SwitchIO70313.xExitEnable:=(ConveyorIO70199.xEmpty AND (ConveyorIO70152.diDesConveyor=70199 OR ConveyorIO70152.diDesConveyor=70154))
													OR (ConveyorIO701100.xEmpty AND (ConveyorIO70152.diDesConveyor=701100 OR ConveyorIO70152.diDesConveyor=70155));
ConveyorIO70192.xUnloadCCW:=ConveyorIO70192.diDesConveyor=701100 OR ConveyorIO70192.diDesConveyor=70155;
ConveyorIO70199.xLoad:=ConveyorIO70192.xNextRun AND (ConveyorIO70152.diDesConveyor=70199 OR ConveyorIO70152.diDesConveyor=70154);
ConveyorIO70199.xUnload:=ConveyorIO70154.xEmpty AND ConveyorIO70199.diDesConveyor=70154;
ConveyorIO70154.xLoad:=ConveyorIO70199.xNextRun;
m_xtonConveyor70199Reset(IN:=NOT ConveyorIO70199.xCWPresent,PT:=T#10s ,Q:= ConveyorIO70199.xPutInto,ET:= m_xtonConveyor70199CurTime );
m_xtonConveyor70154Reset(IN:=NOT ConveyorIO70154.xCWPresent,PT:=T#10s ,Q:= ConveyorIO70154.xPutInto,ET:= m_xtonConveyor70154CurTime );
ConveyorIO701100.xLoad:=ConveyorIO70192.xNextRun AND (ConveyorIO70152.diDesConveyor=701100 OR ConveyorIO70152.diDesConveyor=70155);
ConveyorIO701100.xUnload:=ConveyorIO70155.xEmpty AND ConveyorIO701100.diDesConveyor=70155;
ConveyorIO70155.xLoad:=ConveyorIO701100.xNextRun;
m_xtonConveyor701100Reset(IN:=NOT ConveyorIO701100.xCWPresent,PT:=T#10s ,Q:= ConveyorIO701100.xPutInto,ET:=m_xtonConveyor701100CurTime );
m_xtonConveyor70155Reset(IN:=NOT ConveyorIO70155.xCWPresent,PT:=T#10s ,Q:= ConveyorIO70155.xPutInto,ET:= m_xtonConveyor70155CurTime);



(*3#下层入库*)
(*
IF  ConveyorIO70160.xLoad
	THEN Y2C6:=1;
END_IF;
IF NOT  ConveyorIO70160.xEmpty
	THEN  Y2C6:=0;
END_IF;*)
switch70315(ConveyorEntryIO:= ConveyorIO70160 ,ConveyorExitIO:= ConveyorIO70194 ,SwitchIO:= SwitchIO70315);
SwitchIO70315.xLiftCylinderExtendInit:=1;
SwitchIO70315.xSwithEnable:=1;
Y2C6:=SwitchIO70315.xLiftCylinderExtend;
SwitchIO70315.xLiftCylinderExtendDetect:=XDA;
SwitchIO70315.xLiftCylinderRetractDetect:=XDB;

SwitchIO70315.xExitEnable:=(ConveyorIO701103.xEmpty AND (ConveyorIO70160.diDesConveyor=701103 OR ConveyorIO70160.diDesConveyor=70162))
													OR (ConveyorIO701104.xEmpty AND (ConveyorIO70160.diDesConveyor=701104 OR ConveyorIO70160.diDesConveyor=70163));
ConveyorIO70194.xUnloadCCW:=ConveyorIO70194.diDesConveyor=701103 OR ConveyorIO70194.diDesConveyor=70162;
ConveyorIO701103.xLoad:=ConveyorIO70194.xNextRun AND (ConveyorIO70160.diDesConveyor=701103 OR ConveyorIO70160.diDesConveyor=70162);
ConveyorIO701103.xUnload:=ConveyorIO70162.xEmpty AND ConveyorIO701103.diDesConveyor=70162;
ConveyorIO70162.xLoad:=ConveyorIO701103.xNextRun;
m_xtonConveyor701103Reset(IN:=NOT ConveyorIO701103.xCWPresent,PT:=T#10s ,Q:= ConveyorIO701103.xPutInto,ET:= m_xtonConveyor701103CurTime );
m_xtonConveyor70162Reset(IN:=NOT ConveyorIO70162.xCWPresent,PT:=T#10s ,Q:= ConveyorIO70162.xPutInto,ET:= m_xtonConveyor70162CurTime );
ConveyorIO701104.xLoad:=ConveyorIO70194.xNextRun AND (ConveyorIO70160.diDesConveyor=701104 OR ConveyorIO70160.diDesConveyor=70163);
ConveyorIO701104.xUnload:=ConveyorIO70163.xEmpty AND ConveyorIO701104.diDesConveyor=70163;
ConveyorIO70163.xLoad:=ConveyorIO701104.xNextRun;
m_xtonConveyor701104Reset(IN:=NOT ConveyorIO701104.xCWPresent,PT:=T#10s ,Q:= ConveyorIO701104.xPutInto,ET:=m_xtonConveyor701104CurTime );
m_xtonConveyor70163Reset(IN:=NOT ConveyorIO70163.xCWPresent,PT:=T#10s ,Q:= ConveyorIO70163.xPutInto,ET:= m_xtonConveyor70163CurTime);


(*2，3#下层出库,只写了3#的*)
(*23出库任务抢占*)
	m_Task70314(xCondition:= m_Task70314Condition ,
							xTaskComplete:=LDP(TRUE,ConveyorIO70193.xEmpty) ,
							xReset:= g_xResetSingle AND g_diDeviceIDSelect=70193 ,
							iPriority:= m_iTask70314  );
		m_Task70314Condition[1]:=NOT ConveyorIO701101.xEmpty;
		m_Task70314Condition[2]:=NOT ConveyorIO701102.xEmpty;
		
m_xtonConveyor70159Reset(IN:= ConveyorIO70159.xCWPresent,PT:=T#10s ,Q:= ConveyorIO70159.xPutInto,ET:= m_xtonConveyor70159CurTime );
m_xtonConveyor701102Reset(IN:= ConveyorIO701102.xCWPresent,PT:=T#10s ,Q:= ConveyorIO701102.xPutInto,ET:= m_xtonConveyor701102CurTime );
ConveyorIO70159.xUnload:=ConveyorIO701102.xEmpty;
ConveyorIO701102.xLoad:=ConveyorIO70159.xNextRun;
ConveyorIO701102.xUnload:=ConveyorIO70193.xEmpty AND m_iTask70314=2;

m_xtonConveyor70158Reset(IN:= ConveyorIO70158.xCWPresent,PT:=T#10s ,Q:= ConveyorIO70158.xPutInto,ET:= m_xtonConveyor70158CurTime );
m_xtonConveyor701101Reset(IN:= ConveyorIO701101.xCWPresent,PT:=T#10s ,Q:= ConveyorIO701101.xPutInto,ET:= m_xtonConveyor701101CurTime );
ConveyorIO70158.xUnload:=ConveyorIO701101.xEmpty;
ConveyorIO701101.xLoad:=ConveyorIO70158.xNextRun;
ConveyorIO701101.xUnload:=ConveyorIO70193.xEmpty AND m_iTask70314=1;

ConveyorIO70193.xLoad:=ConveyorIO701102.xNextRun OR ConveyorIO701101.xNextRun;
ConveyorIO70193.xloadCCW:=ConveyorIO701102.xNextRun;
IF  NOT ConveyorIO70193.xEmpty
	THEN Y2C4:=1;(*193转去156顶升*)
END_IF;
ConveyorIO70156.xLoad:= NOT ConveyorIO70193.xEmpty ;
IF NOT  ConveyorIO70156.xEmpty
	THEN 
	Y2C4:=0;
END_IF;
m_xtonConveyor70156Reset(IN:=NOT ConveyorIO70156.xCWPresent,PT:=T#10s ,Q:= ConveyorIO70156.xPutInto,ET:= m_xtonConveyor70156CurTime );
Y33B:=ConveyorIO701102.xNextRun;(*3#出库阻挡*)
Y33A:=ConveyorIO701101.xNextRun;(*2#出库阻挡*)
ConveyorIO70193.xPutInto:=NOT  ConveyorIO70156.xEmpty;
(*最靠近电柜那个出库线体*)
switch70327(ConveyorEntryIO:=ConveyorIO701118,ConveyorExitIO:= ConveyorIO701116_1 ,SwitchIO:= SwitchIO70327);
Y2DE:=SwitchIO70327.xLiftCylinderExtend;
SwitchIO70327.xLiftCylinderExtendDetect:=X155;
SwitchIO70327.xLiftCylinderRetractDetect:=X156;

Conveyor701116_1(ConveyorMotor:= ConveyorIO701116_1 );
ConveyorIO701116_1.xCWPresent:=ConveyorIO701118.xCWPresent;

m_xtonConveyor701120Reset(IN:=ConveyorIO701120.xCWPresent,PT:=T#10s ,Q:= ConveyorIO701120.xPutInto,ET:= m_xtonConveyor701120CurTime );
m_xtonConveyor701119Reset(IN:=ConveyorIO701119.xCWPresent,PT:=T#10s ,Q:= ConveyorIO701119.xPutInto,ET:= m_xtonConveyor701119CurTime );
ConveyorIO701119.tLoadDelay:=t#3s;
ConveyorIO701120.xUnload:=ConveyorIO701119.xEmpty;
ConveyorIO701119.xLoad:=ConveyorIO701120.xNextRun;
ConveyorIO701119.xUnload:=ConveyorIO701118.xEmpty;
SwitchIO70327.xEntryEnable:=ConveyorIO701119.xNextRun;
SwitchIO70327.xSwithEnable:=1;
SwitchIO70327.xExitEnable:=ConveyorIO701116.xEmpty;
ConveyorIO701116.xLoad:=ConveyorIO701116_1.xNextRun;

(*回流部分去分容线体*)
ConveyorIO70141.xLoad:=X3D;
Y2BA:=ConveyorIO70141.xEmpty;
m_xtonConveyor70141Reset(IN:=NOT ConveyorIO70141.xCWPresent,PT:=T#8s ,Q:= ConveyorIO70141.xPutInto,ET:= m_xtonConveyor70141CurTime );

(*————————上层空框回流————————————*)
ConveyorIO70134.xUnload:=ConveyorIO70133.xEmpty;
ConveyorIO70133.xLoad:=ConveyorIO70134.xNextRun;
ConveyorIO70133.xUnload:=ConveyorIO70132.xEmpty;
ConveyorIO70132.xLoad:=ConveyorIO70133.xNextRun;
ConveyorIO70132.xUnload:=ConveyorIO70131.xEmpty;
ConveyorIO70131.xLoad:=ConveyorIO70132.xNextRun;
ConveyorIO70131.xUnload:=ConveyorIO70130.xEmpty;
ConveyorIO70130.xLoad:=ConveyorIO70131.xNextRun;
ConveyorIO70130.xUnload:=ConveyorIO70124.xEmpty;
ConveyorIO70124.xLoad:=ConveyorIO70130.xNextRun;
ConveyorIO70124.xUnload:=ConveyorIO70123.xEmpty;
ConveyorIO70123.xLoad:=ConveyorIO70124.xNextRun;
ConveyorIO70123.xUnload:=ConveyorIO70122.xEmpty;
ConveyorIO70122.xLoad:=ConveyorIO70123.xNextRun;
ConveyorIO70122.xUnload:=ConveyorIO70116.xEmpty;
ConveyorIO70116.xLoad:=ConveyorIO70122.xNextRun;
ConveyorIO70116.xUnload:=ConveyorIO70115.xEmpty;
ConveyorIO70115.xLoad:=ConveyorIO70116.xNextRun;
ConveyorIO70115.xUnload:=ConveyorIO70114.xEmpty;
ConveyorIO70114.xLoad:=ConveyorIO70115.xNextRun;
ConveyorIO70114.xUnload:=ConveyorIO70108.xEmpty;
ConveyorIO70108.xLoad:=ConveyorIO70114.xNextRun;
ConveyorIO70108.xUnload:=ConveyorIO70107.xEmpty AND LifterIO70208.iCurrentPos=2; 
(*提升机2*)
LifterIO70208.xMDIExe:=NOT (ConveyorIO70108.xError OR ConveyorIO70142.xError OR ConveyorIO70107.xError);
IF ConveyorIO70107.xEmpty THEN
	LifterIO70208.iDestinationPos:=2;
ELSE
	LifterIO70208.iDestinationPos:=1;
END_IF;
ConveyorIO70107.xLoad:=ConveyorIO70108.xNextRun AND LifterIO70208.iCurrentPos=2;
ConveyorIO70107.xUnload:=ConveyorIO70142.xEmpty AND  LifterIO70208.iCurrentPos=1;
ConveyorIO70142.xLoad:=ConveyorIO70107.xNextRun AND   LifterIO70208.iCurrentPos=1;







(*临时程序,输送出去,不进2号OCV2，不分拣*) 
(*ConveyorIO70166.xUnload:=ConveyorIO70167.xEmpty;*)
(*临时程序,分拣前顶升移载前*)
(*SwitchIO70319.xEntryEnable:=ConveyorIO70166.xNextRun;*)
(*SwitchIO70319.xSwithEnable:=0;*)(*临时程序不分拣*)
(*SwitchIO70319.xExitEnable:=ConveyorIO70169.xEmpty;
SwitchIO70320.xEntryEnable:=ConveyorIO70167.xNextRun;
SwitchIO70320.xSwithEnable:=1;
SwitchIO70320.xExitEnable:=0;*)(*RGV接料处*)


IF g_xAuto AND NOT g_xRGVTcpFailed THEN
	D201:=m_iRGVDestinationPos;
	D202.0:=g_xRGVRemoteAuto;
	D202.1:=(*ConveyorIO70140.xEmpty*)NOT FolderIO70201.o_xExitPremit;(*更换成叠盘机允许下料信号，RGV生成任务*)
	D202.2:=ConveyorIO701111.xEmpty;
	D202.3:=ConveyorIO70144.xEmpty;
	D202.4:=ConveyorIO70148.xEmpty;
	D202.5:=ConveyorIO70152.xEmpty;
	D202.6:=ConveyorIO70156.xEmpty;
	D202.7:=ConveyorIO70160.xEmpty;
	D202.8:=ConveyorIO70164.xEmpty;
	D202.9:=ConveyorIO70170.xEmpty;
	D202.A:=ConveyorIO70174.xEmpty;
	D202.B:=ConveyorIO701116.xEmpty;
	D203.0:=m_xRGVReset;
	D203.1:=ConveyorIO70140.xNextRun;
	D203.2:=ConveyorIO701111.xNextRun;
	D203.3:=ConveyorIO70148.xNextRun;
	D203.4:=ConveyorIO70156.xNextRun;
	D203.5:=ConveyorIO70170.xNextRun;
	D203.6:=ConveyorIO701116.xNextRun;
	D203.A:=g_SemiStart;
	m_iRGVCurrentPos:=D401;
	m_xRGVPositionArrive:=D401.0;
	m_xRGVConveyorEmpty:=D401.1;
	m_xRGVConveyorNextRun:=D402.2;
	ConveyorIO70140.xUnload:=D402.3;
	ConveyorIO701111.xUnload:=D402.4;
	ConveyorIO70144.xLoad:=D402.5;
	ConveyorIO70148.xUnload:=D402.6;
	ConveyorIO70152.xLoad:=D402.7;
	ConveyorIO70156.xUnload:=D402.8;
	ConveyorIO70160.xLoad:=D402.9;
	ConveyorIO70164.xLoad:=D402.A;
	ConveyorIO70170.xUnload:=D402.B;
	ConveyorIO70174.xLoad:=D402.C;
	ConveyorIO701116.xUnload:=D402.D;
	m_xRGVAlarm:=D403.0;
ELSE
	D201:=0;
	D202:=0;
	D203.0:=0;
	D203.1:=0;
	D203.2:=0;
	D203.3:=0;
	D203.4:=0;
	D203.5:=0;
	ConveyorIO70140.xUnload:=0;
	ConveyorIO701111.xUnload:=0;
	ConveyorIO70144.xLoad:=0;
	ConveyorIO70148.xUnload:=0;
	ConveyorIO70152.xLoad:=0;
	ConveyorIO70156.xUnload:=0;
	ConveyorIO70160.xLoad:=0;
	ConveyorIO70164.xLoad:=0;
	ConveyorIO70170.xUnload:=0;
	ConveyorIO70174.xLoad:=0;
END_IF;
g_xAlarm:=ComConveyorIO70104.i_iResponsPCPLC=101;
END_PROGRAM

FUNCTION_BLOCK PreemptivePriority
VAR_INPUT
  xCondition : ARRAY [1..13] OF BOOL;  (* 条件1 *)
  xTaskComplete : BOOL;  (* 任务完成 *)
  xReset : BOOL;  (* 复位 *)
END_VAR
VAR
  xOccupy : BOOL;  (* 占用 *)
END_VAR
VAR_OUTPUT
  iPriority : INT;  (* 输出任务号 *)
END_VAR
VAR
  m_tonConditionDelay : TON;
  m_xConditionDelay : BOOL;
  m_tConditionCurrentTime : TIME;
  m_iLastTask : INT;  (* 上次执行的任务 *)
  m_tpLastTaskPulse1 : TP;
  m_tpLastTaskPulse2 : TP;
  m_tpLastTaskPulse3 : TP;
  m_tpLastTaskPulse4 : TP;
  m_tpLastTaskPulse5 : TP;
  m_xLastTaskPulse : ARRAY [1..13] OF BOOL;
  m_tLastTaskPulse : ARRAY [1..13] OF TIME := [13(T#0s)];
  m_tpLastTaskPulse6 : TON;
  ii : INT;
END_VAR
VAR CONSTANT
  CONDITION_QUANTITY : INT := 9;
END_VAR
VAR
  m_tpLastTaskPulse7 : TON;
  m_tpLastTaskPulse8 : TON;
  m_tpLastTaskPulse9 : TON;
  m_tpLastTaskPulse10 : TON;
  m_tpLastTaskPulse11 : TON;
  m_tpLastTaskPulse12 : TON;
  m_tpLastTaskPulse13 : TON;
END_VAR
(*抢占式优先级块
现在满足13个条件的任务进行抢占式优先级排列
条件满足后延时两秒，开始执行任务，
同一任务连续执行优先级下降
需要改造成任意多个
使用于一个入口多个出口的程序，使用抢占式优先级块
*)
IF LDP(TRUE, xTaskComplete) THEN
	xOccupy:=0;
	iPriority:=0;
END_IF;
(*//任务滤波，延时两秒*)
m_tonConditionDelay(IN:=( xCondition[1]
 	OR xCondition[2]
 	OR xCondition[3]
 	OR xCondition[4]
 	OR xCondition[5]
 	OR xCondition[6]
 	OR xCondition[7]
 	OR xCondition[8]
 	OR xCondition[9]
 	OR xCondition[10]
 	OR xCondition[11]
 	OR xCondition[12]
 	OR xCondition[13]
 	)
 	AND iPriority=0,
 PT:= T#1s,
 Q:= m_xConditionDelay ,
 ET:= m_tConditionCurrentTime );		
(*//判断优先级，上个任务与本次任务相同，延时一秒执行*)
m_tpLastTaskPulse1(IN:= xCondition[1]  AND m_iLastTask=1 AND m_xConditionDelay  ,PT:= T#1s,Q:= m_xLastTaskPulse[1],ET:= m_tLastTaskPulse[1] );
m_tpLastTaskPulse2(IN:= xCondition[2]  AND m_iLastTask=2 AND m_xConditionDelay  ,PT:= T#1s,Q:= m_xLastTaskPulse[2],ET:= m_tLastTaskPulse[2] );
m_tpLastTaskPulse3(IN:= xCondition[3]  AND m_iLastTask=3 AND m_xConditionDelay  ,PT:= T#1s,Q:= m_xLastTaskPulse[3],ET:= m_tLastTaskPulse[3] );
m_tpLastTaskPulse4(IN:= xCondition[4]  AND m_iLastTask=4 AND m_xConditionDelay  ,PT:= T#1s,Q:= m_xLastTaskPulse[4],ET:= m_tLastTaskPulse[4] );
m_tpLastTaskPulse5(IN:= xCondition[5]  AND m_iLastTask=5 AND m_xConditionDelay  ,PT:= T#1s,Q:= m_xLastTaskPulse[5],ET:= m_tLastTaskPulse[5] );
m_tpLastTaskPulse6(IN:= xCondition[6]  AND m_iLastTask=6 AND m_xConditionDelay  ,PT:= T#1s,Q:= m_xLastTaskPulse[6],ET:= m_tLastTaskPulse[6] );
m_tpLastTaskPulse7(IN:= xCondition[7]  AND m_iLastTask=7 AND m_xConditionDelay  ,PT:= T#1s,Q:= m_xLastTaskPulse[7],ET:= m_tLastTaskPulse[7] );
m_tpLastTaskPulse8(IN:= xCondition[8]  AND m_iLastTask=8 AND m_xConditionDelay  ,PT:= T#1s,Q:= m_xLastTaskPulse[8],ET:= m_tLastTaskPulse[8] );
m_tpLastTaskPulse9(IN:= xCondition[9]  AND m_iLastTask=9 AND m_xConditionDelay  ,PT:= T#1s,Q:= m_xLastTaskPulse[9],ET:= m_tLastTaskPulse[9] );
m_tpLastTaskPulse10(IN:= xCondition[10]  AND m_iLastTask=10 AND m_xConditionDelay  ,PT:= T#1s,Q:= m_xLastTaskPulse[10],ET:= m_tLastTaskPulse[10] );
m_tpLastTaskPulse11(IN:= xCondition[11]  AND m_iLastTask=11 AND m_xConditionDelay  ,PT:= T#1s,Q:= m_xLastTaskPulse[11],ET:= m_tLastTaskPulse[11] );
m_tpLastTaskPulse12(IN:= xCondition[12]  AND m_iLastTask=12 AND m_xConditionDelay  ,PT:= T#1s,Q:= m_xLastTaskPulse[12],ET:= m_tLastTaskPulse[12] );
m_tpLastTaskPulse13(IN:= xCondition[13]  AND m_iLastTask=13 AND m_xConditionDelay  ,PT:= T#1s,Q:= m_xLastTaskPulse[13],ET:= m_tLastTaskPulse[13] );
(*//执行*)
FOR ii:=1 TO CONDITION_QUANTITY BY 1 DO 
	IF NOT xCondition[ii] AND NOT xOccupy THEN
		iPriority:=0;
	END_IF;
	IF xCondition[ii] AND NOT xOccupy AND m_xConditionDelay AND NOT  m_xLastTaskPulse[ii]  THEN
		iPriority:=ii;
		xOccupy:=1;
		m_iLastTask:=ii;
	END_IF;
END_FOR;        
(*//复位*)
IF xReset THEN
	iPriority:=0;
	xOccupy:=0;
	m_iLastTask:=0;	
END_IF;
(*//清除占用*)
IF iPriority=0 THEN
	xOccupy:=0;
END_IF;
END_FUNCTION_BLOCK

FUNCTION_BLOCK PriorityQueue
VAR_INPUT
  arrxCondition : ARRAY [1..13] OF QueueElement;
  xTaskComplete : BOOL;  (* 任务完成 *)
  xReset : BOOL;  (* 复位 *)
END_VAR
VAR
  xOccupy : BOOL;  (* 占用 *)
END_VAR
VAR_OUTPUT
  iPriority : INT;  (* 输出任务号 *)
END_VAR
VAR
  jj : INT;
END_VAR
VAR CONSTANT
  CONDITION_QUANTITY : INT := 9;
END_VAR
VAR_IN_OUT
  arriTaskStack : ARRAY [0..13] OF INT;
END_VAR
VAR
  ii : INT;
  kk : INT;
  arrxConditionDelay : ARRAY [1..13] OF BOOL;
  arrxConditionEdgeDetect : ARRAY [1..13] OF BOOL;
  arrxDelayEdgeDetect : ARRAY [1..13] OF BOOL;
  arriDelayCounter : ARRAY [1..13] OF INT;
  ll : INT;
  Temp : INT;
  mm : INT;
  nn : INT;
  Temp2 : INT;
  oo : INT;
END_VAR
(****************************************************************************)
(*
一般情况多对一的任务调度采用这个结构，排队通过出口
优先级功能块，存储任意条件的优先级，实现栈功能先入先出，
复位功能还有问题，
出入栈式优先级块，满足条件后入栈，先入先出，在栈尾加载新任务
栈首为当前执行的任务，任务完成使用上升沿触发，触发后栈首元素弹出

复位功能清空堆栈，栈的容量在CONDITION_QUANTITY 设置
增加了结构体，结构体中带有一个条件函数，和一个优先级指示
任务完成后通过凭借优先级来排序，优先级高的条件先执行   优先级排序是从小到大的，数值小的优先级高
防止干扰，增加了任务的1秒的延时
*)

(***************************************************************************)
(*(//入栈*)
FOR ii:=1 TO CONDITION_QUANTITY BY 1 DO
	(*//循环内无法用定时器，改用计数器的形式*)
	IF arrxCondition[ii].xCondition AND SM411 (*//0.2秒的方波信号，如果移植需要修改成两个定时器*)
		AND arriDelayCounter[ii]<6  (* //计数为6，5个0.2秒的方波，所以为1秒*)
		AND NOT arrxDelayEdgeDetect[ii] THEN    (*//循环内无法用沿函数，增加锁定标志位*)
		arriDelayCounter[ii]:=arriDelayCounter[ii]+1;   (*//计数*)
	END_IF;
	IF NOT arrxCondition[ii].xCondition THEN
		arriDelayCounter[ii]:=0;   (*//计数清零*)
	END_IF;
	arrxDelayEdgeDetect[ii]:=arrxCondition[ii].xCondition AND SM411;  (*//沿函数锁*)
	IF arriDelayCounter[ii]=5 AND NOT arrxConditionEdgeDetect[ii] THEN;  (*//条件满足1秒后*)
		FOR kk:=0 TO CONDITION_QUANTITY BY 1 DO    
			IF arriTaskStack[kk]=0 THEN
				arriTaskStack[kk]:=ii;   (*//栈尾添加*)
				EXIT;
			END_IF;		
		END_FOR;
	END_IF;	
	arrxConditionEdgeDetect[ii]:=arriDelayCounter[ii]=5;  (*//边沿*)
END_FOR;
(*//栈顶任务为当前执行的任务**)
iPriority:=arriTaskStack[0]; 
(*//栈顶任务完成，弹出*)
IF 	LDP(TRUE, xTaskComplete) THEN
	FOR jj:=0 TO CONDITION_QUANTITY-1 BY 1 DO
		arriTaskStack[jj]:=arriTaskStack[jj+1];
	END_FOR;
	arriTaskStack[CONDITION_QUANTITY]:=0;(*//栈尾清零*)
	(*//排序，使用插入排序*)
	FOR oo:=0 TO CONDITION_QUANTITY BY 1 DO
		IF arriTaskStack[oo]=0 THEN
			EXIT;  (* //寻找栈中不为零的元素  ，防止0元素进入条件查找的时候报错*)
		END_IF;
	END_FOR;
	(*//插入排序insertionsort*)
	FOR mm:=1 TO oo-1  BY 1 DO   (*//从1开始*)
		Temp:=arriTaskStack[mm];  (*//当前数据记录 *)
		Temp2:=arrxCondition[arriTaskStack[mm]].iPriority;  (*//当前优先级记录 *)
		nn:=mm;  (*//指针赋值*)
		WHILE  (nn>0 AND Temp2< arrxCondition[arriTaskStack[nn-1]].iPriority)  DO  (*//优先级比较，当前优先级小于他前面元素优先级的时候*)
			 arriTaskStack[nn] := arriTaskStack[nn-1] ;  (*//优先级低的向后复制，比TEMP2大的元素都要复制到下一个位置*)
			 nn:=nn-1;
		END_WHILE;
		arriTaskStack[nn]:=Temp; (*//把当前数据放在合适的位置*)
	END_FOR;
END_IF;
(*//复位*)
IF xReset THEN
	FOR jj:=0 TO CONDITION_QUANTITY BY 1 DO
		arriTaskStack[jj]:=0;
	END_FOR;
	FOR ll:=1 TO CONDITION_QUANTITY BY 1 DO
		arrxConditionEdgeDetect[ll]:=0;
		arriDelayCounter[ll]:=0;
	END_FOR;
END_IF;
END_FUNCTION_BLOCK

FUNCTION_BLOCK Servo
Y380:=1;
END_FUNCTION_BLOCK

FUNCTION_BLOCK ShuttleCar
VAR_IN_OUT
  ShuttleCarInOut : ShuttleCarIO;
END_VAR
VAR
  m_tonBrakeDelay : TON;  (* 延时 *)
  m_tBrakeDelayCurrentTime : TIME;
  m_tonArriveDelay : TON;  (* 到达延时计时器 *)
  m_xArriveDelay : BOOL;  (* 到达延时 *)
  m_tArriveDelayCurrentTime : TIME;  (* 到达延时当前时间 *)
  m_xInit : BOOL;  (* 初始化标志位 *)
  m_tonPauseDelay : TON;  (* 暂停减速 *)
  m_tPauseDelayCurrentTime : TIME;  (* 暂停延时当前时间 *)
  m_tonOvertimeAlarm : TON;  (* 超时报警定时器 *)
  m_tOvertimeCurrentTime : TIME;  (* 超时报警当前时间 *)
END_VAR
(*******************************************************************
输送小车程序，可用于使用认址片控制位置的输送车程序，可用于控制提升机，
使用了限位捕捉程序防止小车惯性过大冲过限位后继续行走，捕捉程序采用反
转复位，这样设计有弊端可能反转复位后车的位置并没有回到限位以内,当两个
限位同时碰到的时候，会使运料小车进入死锁状态，通过xPassLimit来解开死锁，
可以在触摸屏中使用一个带权限的按钮来进行控制，配合ShuttleCarCurrentPos
函数来计算位置信息
增加自动开始后将当前位置置为零的信号防止设备停在两个位置开关的中间
修改信息  修改后请增加版本
2018-1-22增加到位延时：到位延时时间可以设置，适应双向到位的位置开关，通过调整延时时间让穿梭车停在到位开关的中间
增加气缸控制信号 ShuttleCarInOut.xCylinder
增加抱闸延时 ShuttleCarInOut.tBrakeDelay
增加超时报警 ShuttleCarInOut.xOvertimeAlarm
YAO      V1.0
2018-1-22 YAO V1.1
2018-6-3：增加点动xMoveStep，单体报警复位
接口说明：
输入：
xReady    准备就绪信号，接变频器的准备就绪，无准备就绪信号的设备常置1
xForward   手动 正转
xBackward 手动 反转
iCurrentPos 当前位置信息，由外部函数给出
iDestinationPos  目标位置，自动情况下判断目标位置和当前位置的差，选择前进或后退
xPosLimit 正方向限位  常闭信号
xNegLimit 反方向限位  常闭信号
xMDIExe   自动行走使能
xPassLimit 限位屏蔽
tArriveDelay 到位延时时间设置，当前位置等于目标位置后延时相应时间后停止，默认为0
xCylinder 如果是气缸的把这个标志位置为1，
tBrakeDelay 打开抱闸延时，默认100ms。行走后会延时相应的时间打开抱闸，防止提升轴的掉落
xLooseDetect 松绳检测开关
输出：
xCW 正转输出
xCCW 反转输出
xBrake 抱闸输出 
xMDIDone 自动行走完成信号
xPosLimitCatch 正限位报警
xNegLimitCatch 负限位报警
xBusy 工作中信号
xLooseAlarm 松绳报警，报警后不可以下降，提升后如果没有松绳检测开关后复位报警信号


********************************************************************)
IF NOT m_xInit THEN
	ShuttleCarInOut.tArriveDelay:=T#0s;   (*到位延时初始化为0*)
	ShuttleCarInOut.tBrakeDelay:=T#100ms;(*抱闸延时初始化为100ms*)
	ShuttleCarInOut.tSetOverTime:=T#60s;(*超时报警初始化为1分钟*)
	m_xInit:=1;
END_IF;
(*如果是气缸的话屏蔽限位和Ready信号*)
IF ShuttleCarInOut.xCylinder THEN
	ShuttleCarInOut.xPosLimit:=1;
	ShuttleCarInOut.xNegLimit:=1;
	ShuttleCarInOut.xReady:=1;
END_IF;
(*限位捕捉，防止冲过限位开关，反转后复位*)
ShuttleCarInOut.xPosLimitCatch:=LDF(TRUE,ShuttleCarInOut.xPosLimit) OR ShuttleCarInOut.xPosLimitCatch;
IF ShuttleCarInOut.xCCW THEN  
	ShuttleCarInOut.xPosLimitCatch:=0;
END_IF;

ShuttleCarInOut.xNegLimitCatch:=LDF(TRUE,ShuttleCarInOut.xNegLimit) OR ShuttleCarInOut.xNegLimitCatch;
(*松绳报警*)
IF LDP(TRUE,ShuttleCarInOut.xLooseDetect) THEN	
	ShuttleCarInOut.xLooseAlarm:=1;
END_IF;
(*提升复位报警*)
IF ShuttleCarInOut.xCW AND NOT  ShuttleCarInOut.xLooseDetect THEN   
	ShuttleCarInOut.xLooseAlarm:=0; 
END_IF;

IF ShuttleCarInOut.xCW THEN   
	ShuttleCarInOut.xNegLimitCatch:=0; 
END_IF;

IF ShuttleCarInOut.xPassLimit OR
	g_xReset OR   (*增加复位按钮*)
	(ShuttleCarInOut.xNegLimitCatch 
	AND ShuttleCarInOut.xPosLimitCatch)  THEN  
	ShuttleCarInOut.xNegLimitCatch:=0; 
	ShuttleCarInOut.xPosLimitCatch:=0;
	ShuttleCarInOut.xLooseAlarm:=0;
END_IF;
IF ShuttleCarInOut.xReady AND g_xEStop THEN
(*手动*)
    IF g_xManual THEN  
	    IF ShuttleCarInOut.xForward 
			AND ShuttleCarInOut.xBackward=0 
			AND ShuttleCarInOut.xCCW=0 
			AND ShuttleCarInOut.xPosLimitCatch=0  THEN
		    ShuttleCarInOut.xCW:=1;
		    ELSE
		    ShuttleCarInOut.xCW:=0;
	    END_IF;
	    IF ShuttleCarInOut.xBackward 
			AND ShuttleCarInOut.xForward=0 
			AND ShuttleCarInOut.xCW=0 
			AND ShuttleCarInOut.xNegLimitCatch=0 
			AND ShuttleCarInOut.xLooseAlarm=0
			AND G_xEStop THEN  
		    ShuttleCarInOut.xCCW:=1;
		    ELSE
		    ShuttleCarInOut.xCCW:=0;
	    END_IF;
    END_IF;
    (**********)
(*自动*)
  IF g_xAuto OR ShuttleCarInOut.xMoveStep   THEN  
  	(*点动*)
  	IF LDP(TRUE,ShuttleCarInOut.xMoveStep)  THEN (*点动模式后把当前位置赋值给目标位置，防止误动作*)
  		ShuttleCarInOut.iDestinationPos:=ShuttleCarInOut.iCurrentPos;
  		END_IF;
 		IF LDP(TRUE,ShuttleCarInOut.xForward) AND ShuttleCarInOut.xMoveStep THEN
 			ShuttleCarInOut.xMDIExe:=1;
			ShuttleCarInOut.iDestinationPos:=ShuttleCarInOut.iCurrentPos+1;
		END_IF;
		IF LDP(TRUE,ShuttleCarInOut.xBackward) AND ShuttleCarInOut.xMoveStep AND ShuttleCarInOut.iCurrentPos>0  THEN
			ShuttleCarInOut.xMDIExe:=1;
			ShuttleCarInOut.iDestinationPos:=ShuttleCarInOut.iCurrentPos-1;
		END_IF;	 
	(*>>>>>>>>>>>>>>>>>>>>>>>>>>>>>>>>>>>>>*)	
	  IF ShuttleCarInOut.xMDIExe AND ShuttleCarInOut.iDestinationPos<>0 THEN	
	    IF ShuttleCarInOut.iCurrentPos<ShuttleCarInOut.iDestinationPos AND ShuttleCarInOut.xPosLimitCatch=0 THEN   (*正转*)
			ShuttleCarInOut.xCW:=1;
			ShuttleCarInOut.xCCW:=0;
			ShuttleCarInOut.xMDIDone:=0;
		END_IF;

		IF ShuttleCarInOut.iCurrentPos>ShuttleCarInOut.iDestinationPos AND ShuttleCarInOut.xNegLimitCatch=0 AND ShuttleCarInOut.xLooseAlarm=0 THEN   (*反转*)
			ShuttleCarInOut.xCCW:=1;
			ShuttleCarInOut.xCW:=0;
			ShuttleCarInOut.xMDIDone:=0;
		END_IF;
	m_tonArriveDelay(IN:= ShuttleCarInOut.iCurrentPos=ShuttleCarInOut.iDestinationPos ,
	                                    PT:= ShuttleCarInOut.tArriveDelay ,
	                                    Q:= m_xArriveDelay ,
	                                    ET:= m_tArriveDelayCurrentTime);
	     (*到位延时时间可以设置，适应双向到位的位置开关，通过调整延时时间让穿梭车停在到位开关的中间*)
		IF m_xArriveDelay AND NOT ShuttleCarInOut.xCylinder THEN
			ShuttleCarInOut.xCW:=0;
			ShuttleCarInOut.xCCW:=0;
			ShuttleCarInOut.xMDIDone:=1;
			ELSE
			ShuttleCarInOut.xMDIDone:=0;
		END_IF;

		IF ShuttleCarInOut.xPosLimitCatch THEN
			ShuttleCarInOut.xCW:=0;
			ShuttleCarInOut.xMDIDone:=0;
		END_IF;

		IF ShuttleCarInOut.xNegLimitCatch  OR ShuttleCarInOut.xLooseAlarm THEN
			ShuttleCarInOut.xCCW:=0;
			ShuttleCarInOut.xMDIDone:=0;
		END_IF;
		ELSE
		ShuttleCarInOut.xCW:=0;
		ShuttleCarInOut.xCCW:=0;
		ShuttleCarInOut.xMDIDone:=0;
	  END_IF;
	END_IF;
	ELSE  (*无就绪信号   或急停的情况下*)
		ShuttleCarInOut.xCW:=0;
		ShuttleCarInOut.xCCW:=0;	
END_IF;
    (*抱闸延时*)
m_tonBrakeDelay(IN:= ShuttleCarInOut.xCW OR ShuttleCarInOut.xCCW,
                                    PT:= ShuttleCarInOut.tBrakeDelay,
                                    Q:=ShuttleCarInOut.xBrake ,
                                    ET:= m_tBrakeDelayCurrentTime);

(*自动上电后把当前位置清零，防止穿梭车不在开关位置*)
IF LDP(TRUE,g_xAuto) THEN
	ShuttleCarInOut.iCurrentPos:=0;
END_IF;
IF ShuttleCarInOut.xCW OR ShuttleCarInOut.xCCW THEN
	ShuttleCarInOut.xBusy:=1;
	ELSE
	ShuttleCarInout.xBusy:=0;
END_IF;

(*暂停，带延时减速斜坡，ShuttleCarInOut.xPauseRamp为减速斜坡输出位*)
m_tonPauseDelay(IN:=g_xPause,PT:= T#2s ,Q:=ShuttleCarInOut.xPauseRamp,ET:= m_tPauseDelayCurrentTime );
IF ShuttleCarInOut.xPauseRamp THEN
	ShuttleCarInOut.xCW:=0;
	ShuttleCarInOut.xCCW:=0;
	ShuttleCarInOut.xBrake:=0;
END_IF;
(*超时报警*)
m_tonOvertimeAlarm(IN:= ShuttleCarInOut.xMDIExe AND (ShuttleCarInOut.iCurrentPos<>ShuttleCarInOut.iDestinationPos) ,
                                           PT:= ShuttleCarInOut.tSetOverTime,
                                           Q:= ShuttleCarInOut.xOvertimeAlarm ,
                                           ET:= m_tOvertimeCurrentTime );
(*//单体复位，当设备号与本设备一致的时候执行复位*)
IF (g_xResetSingle AND ShuttleCarInOut.diDeviceID=g_diDeviceIDSelect)THEN(*增加单体复位*)
	ShuttleCarInOut.iCurrentPos:=0;
END_IF;
END_FUNCTION_BLOCK

FUNCTION ShuttleCarCurrentPosition
VAR_INPUT
  xPosition1 : BOOL;
  xPosition2 : BOOL;
  xPosition3 : BOOL;
END_VAR
(*//计算输送车当前位置的函数*)
IF xPosition1 THEN
	ShuttleCarCurrentPosition:=1;
END_IF;
IF xPosition2 THEN
	ShuttleCarCurrentPosition:=2;
END_IF;
IF xPosition3 THEN
	ShuttleCarCurrentPosition:=3;
END_IF;
END_FUNCTION

FUNCTION_BLOCK SortCommunication
VAR
  m_iStep : INT;
END_VAR
VAR_IN_OUT
  ConveyorIO : ConveyorIO;
  SortCommunicationIO : SortCommunicationIO;
END_VAR
VAR
  m_iCoordinateX : INT;
  m_iCoordinateY : INT;
END_VAR
VAR_IN_OUT
  FanucRobotIO : FanucRobotIO;
END_VAR
VAR_OUTPUT
  o_iErrorNub : INT;
END_VAR
VAR
  ii : INT;
END_VAR
VAR CONSTANT
  ROW_NUB : INT := 8;  (* 每排的数量 *)
END_VAR
VAR
  m_xEno : BOOL;
  m_TONPutover : TON;  (* 放货完成滤波 *)
  m_xPutover : BOOL;  (* 放货完成滤波 *)
  m_tPutover : TIME;  (* 放货完成滤波 *)
  m_iCheck : INT;  (* 校验字 *)
END_VAR
(*********************************************************)
(*
DB1区(PC->PLC)100个字		
"字(16位）序号
(从1开始)"	功能描述	具体参数解释
1	应答	"1：复位
2：读码成功(参数写入完成)
101：条码空
102：条码规则校验失败
103：步号校验失败"
2	任务处理完成	"1：复位
2：处理完成"
3	"电芯状态，
128个电芯"	一个字代表两个电芯状态，1：合格，2,3,4:NG 

DB2区(PLC->PC)10个字		
"字(16位）序号
(从1开始)"	功能描述	具体参数解释
请求	"1：无板
2：请求分拣
"
分拣完成	"1：复位
2：挑选完成
3：撤销
"
跟机器人通信13个输出，2个输入
						13个输出分别是：4个表示行，4个表示列，4个表示不良信息，1个启动信号
						2个输入分别是：抓料完成，放料完成		

*)
(*********************************************************)
IF g_xAuto THEN
	(*——这里临时改一下，暂时人工挑选,所以需要分拣完成按钮——*)	
		IF LDP(TRUE,SortCommunicationIO.i_xSortOver)THEN
			m_iStep:=4;
		END_IF;(**)
		(*夹紧气缸控制*)
		FanucRobotIO.o_xCatchCylinder:=NOT  ConveyorIO.xEmpty AND NOT SortCommunicationIO.o_xSortDone;
		
(*——以上是暂时人工分拣的，以后删掉——*)
	CASE m_iStep OF
		0:(*//初始化*)
		SortCommunicationIO.o_iRequestPLCPC:=1;
		SortCommunicationIO.o_iSortDonePLCPC:=1;
		ii:=0;
		SortCommunicationIO.o_xSortDone:=0;
		m_iStep:=1;
		
		1:(*发送框码的扫码请求*)
		IF ConveyorIO.xEmpty THEN
			SortCommunicationIO.o_iRequestPLCPC:=1;
		ELSE
			SortCommunicationIO.o_iRequestPLCPC:=2;(*发2表示有料了，他就会扫码*)
		END_IF;
		(*//请求确认*)
		IF SortCommunicationIO.o_iRequestPLCPC=2 THEN(*加个条件，免得无脑跳Step2*)
			CASE SortCommunicationIO.i_iResponsPCPLC OF 
			0:;
			1:;(*//复位*)
			2:(*//读码（入库申请）成功*)
				m_iStep:=2;
				ii:=0;
				m_iCoordinateX:=1;(*//框码扫码成功后把坐标改为1,1*)
				m_iCoordinateY:=1;
			3:(*//取放货完成*)
				ConveyorIO.xPutInto:=1; 
			4:(*//旋转*)
				;
			5:(*//不旋转*)
				;
			101:(*//条码空*)
				o_iErrorNub:=101;
			102:(*//条码规则检验失败*)
				o_iErrorNub:=102;
			103:(*//步号校验失败*)
				o_iErrorNub:=103;
			104:(*//无库位可用*)
				o_iErrorNub:=104;
			END_CASE;
		END_IF;	